   M30xTrimDeck_xOSR_OpenOnCleaning : BOOL; {access Read Only}
   M30xTrimDeckAutoResetOppOpSide : TIMER[5] := ([0].PRE := 500); {access Read Only}
   M30xTrimDeckAutoResetOppOpSideTimeout : TIMER[5] := ([0].PRE := 2000); {access Read Only}
   M30xTrimDeckAutoResetOpSide : TIMER[5] := ([0].PRE := 500); {access Read Only}
   M30xTrimDeckAutoResetOpSideTimeout : TIMER[5] := ([0].PRE := 2000); {access Read Only}
   M30xTrimDeckDriveErrorOppOpSide : TIMER[5] := ([0].PRE := 800); {access Read Only}
   M30xTrimDeckDriveErrorOpSide : TIMER[5] := ([0].PRE := 800); {access Read Only}
   M30xTrimWheel : MAC_TrimmingWheels[5] := ([0].CONF_dTrimWheelCodeOpt := 1, [0].CONF_dPositionWheel_cmm := 687500, [0].CONF_dConveyorLength_cmm := 914500, [0].CONF_dMaxLengthWorkable_cmm := 610000, [0].CONF_dTolerance_cmm[0] := 200, [0].CONF_dTolerance_cmm[1] := 200, [0].CONF_dTrimWheelArmPos_cmm[0] := 687500, [0].CONF_dTrimWheelArmPos_cmm[1] := 687500, [0].CONF_dMaxTimeToReachPosition_ms[0] := 600, [0].CONF_dMaxTimeToReachPosition_ms[1] := 600, [0].CONF_dTrimWheelPresetZero_cmm[0] := 2620, [0].CONF_dTrimWheelPresetZero_cmm[1] := 2560, [0].CONF_dTrimWheelTargetWindow_cmm[0] := 200, [0].CONF_dTrimWheelTargetWindow_cmm[1] := 200, [0].CONF_dTrimWheelMinPos_cmm[0] := 115000, [0].CONF_dTrimWheelMinPos_cmm[1] := 115000, [0].CONF_dTrimWheelMaxPos_cmm[0] := 262000, [0].CONF_dTrimWheelMaxPos_cmm[1] := 256000, [0].CONF_dTrimWheelMinRange_cmm[0] := 115000, [0].CONF_dTrimWheelMinRange_cmm[1] := 115000, [0].CONF_dTrimWheelMaxRange_cmm[0] := 262000, [0].CONF_dTrimWheelMaxRange_cmm[1] := 256000, [0].CONF_dAutoSpeed_mm_min[0] := 1000, [0].CONF_dAutoSpeed_mm_min[1] := 1000, [0].CONF_dManualSpeed_mm_min[0] := 200, [0].CONF_dManualSpeed_mm_min[1] := 200, [0].CONF_rAcceleration_m_s2[0] := 1.0, [0].CONF_rAcceleration_m_s2[1] := 1.0, [0].CONF_rDeceleration_m_s2[0] := 1.0, [0].CONF_rDeceleration_m_s2[1] := 1.0, [0].ST_xInitialConditionOpSideOK := 1, [0].ST_xInitialConditionOppOpSideOK := 1, [0].ST_xCleaningConditionOK := 1, [0].ST_xConditionOKStopCycle := 1, [0].ST_xOutputEnableOpSide := 1, [0].ST_xOutputEnableOppOpSide := 1, [0].ST_xEnableControlError := 1, [0].ST_xInPositionOpSide := 1, [0].ST_xInPositionOppOpSide := 1, [0].INPUT_xProtectionMotor := 3, [0].INPUT_xLocalSafetySwitch := 3, [0].INPUT_xMotorThermalProbe := 3, [0].INPUT_xProtectionBrake := 3, [0].INPUT_xBrakeFeedback := 3, [0].INPUT_xDriveReady := 3, [0].INPUT_xHomePosition := 3, [0].OUTPUT_xDriveEnable := 3, [0].AUX_dReqLengthPlate_cmm[0] := 260000, [0].AUX_dReqLengthPlate_cmm[1] := 260000, [0].AUX_dReqPositionPlate_cmm[0] := 965963, [0].AUX_dReqPositionPlate_cmm[1] := 965963, [0].AUX_dReqTargetPosTranslation_cmm[0] := 190430, [0].AUX_dReqTargetPosTranslation_cmm[1] := 186570, [0].AUX_dHeadPosition_cmm[0] := 965963, [0].AUX_dHeadPosition_cmm[1] := 965963, [0].AUX_dLengthPlate_cmm[0] := 260000, [0].AUX_dLengthPlate_cmm[1] := 260000, [0].AUX_dPositionWheelBrk_cmm[0] := 188408, [0].AUX_dPositionWheelBrk_cmm[1] := 187480, [0].AUX_dActTransPosition_cmm[0] := 188408,
        [0].AUX_dActTransPosition_cmm[1] := 187480, [0].AUX_dOffsetStep[0] := 500, [0].AUX_dOffsetStep[1] := 500, [0].AUX_dFinalTarget_cmm[0] := 188430, [0].AUX_dFinalTarget_cmm[1] := 187570, [0].AUX_dReqSpeed_mm_min[0] := 1000, [0].AUX_dReqSpeed_mm_min[1] := 1000, [0].AUX_dRealSpeed_mm_min[0] := 1000, [0].AUX_dRealSpeed_mm_min[1] := 1000, [0].AUX_dTotalCaps[0] := 1, [0].AUX_dTotalCaps[1] := 1, [0].AUX_rgxActivate[0] := 2, [0].AUX_rgxActivate[1] := 2, [0].AUX_dSearchPlateDataOpSide.dReaction_cmm := 1000, [0].AUX_dSearchPlateDataOpSide.dPositionDecision_cmm := 647500, [0].AUX_dSearchPlateDataOpSide.dPositionStopSearch_cmm := 686500, [0].AUX_dSearchPlateDataOpSide.dPositionStopHooked_cmm := 706500, [0].AUX_dSearchPlateDataOppOpSide.dReaction_cmm := 1000, [0].AUX_dSearchPlateDataOppOpSide.dPositionDecision_cmm := 647500, [0].AUX_dSearchPlateDataOppOpSide.dPositionStopSearch_cmm := 686500, [0].AUX_dSearchPlateDataOppOpSide.dPositionStopHooked_cmm := 706500, [0].AUX_dSearchPlateDataTranslationOpSide.dReaction_cmm := 1000, [0].AUX_dSearchPlateDataTranslationOpSide.dPositionDecision_cmm := 647500, [0].AUX_dSearchPlateDataTranslationOpSide.dPositionStopSearch_cmm := 686500, [0].AUX_dSearchPlateDataTranslationOpSide.dPositionStopHooked_cmm := 706500, [0].AUX_dSearchPlateDataTranslationOppOpSide.dReaction_cmm := 1000, [0].AUX_dSearchPlateDataTranslationOppOpSide.dPositionDecision_cmm := 647500, [0].AUX_dSearchPlateDataTranslationOppOpSide.dPositionStopSearch_cmm := 686500, [0].AUX_dSearchPlateDataTranslationOppOpSide.dPositionStopHooked_cmm := 706500, [0].tmON_TrimWheelTimeOut[0].PRE := 2500, [0].tmON_TrimWheelTimeOut[1].PRE := 2500, [0].tmON_TrimWheelBlow[0].PRE := 880, [0].tmON_TrimWheelBlow[0].ACC := 880, [0].tmON_TrimWheelBlow[1].PRE := 800, [0].tmON_TrimWheelBlow[1].ACC := 800, [0].tmOF_DriveEnable[0].PRE := 30000, [0].tmOF_DriveEnable[0].ACC := 9881, [0].tmOF_DriveEnable[0].TT := 1, [0].tmOF_DriveEnable[0].DN := 1, [0].tmOF_DriveEnable[1].PRE := 30000, [0].tmOF_DriveEnable[1].ACC := 9881, [0].tmOF_DriveEnable[1].TT := 1, [0].tmOF_DriveEnable[1].DN := 1, [0].tmON_FeedbackTimeOut[0].PRE := 3500, [0].tmON_FeedbackTimeOut[1].PRE := 3500, [0].tmON_FeedbackDriveReady[0].PRE := 1000, [0].tmON_FeedbackDriveReady[1].PRE := 1000, [1].CONF_dTrimWheelCodeOpt := 2, [1].CONF_dPositionWheel_cmm := 924500, [1].CONF_dConveyorLength_cmm := 914500, [1].CONF_dMaxLengthWorkable_cmm := 610000, [1].CONF_dTolerance_cmm[0] := 200, [1].CONF_dTolerance_cmm[1] := 200, [1].CONF_dTrimWheelArmPos_cmm[0] := 924500, [1].CONF_dTrimWheelArmPos_cmm[1] := 924500, [1].CONF_dMaxTimeToReachPosition_ms[0] := 600, [1].CONF_dMaxTimeToReachPosition_ms[1] := 600, [1].CONF_dTrimWheelPresetZero_cmm[0] := 260, [1].CONF_dTrimWheelPresetZero_cmm[1] := 260, [1].CONF_dTrimWheelTargetWindow_cmm[0] := 200,
        [1].CONF_dTrimWheelTargetWindow_cmm[1] := 200, [1].CONF_dTrimWheelMinPos_cmm[0] := -15000, [1].CONF_dTrimWheelMinPos_cmm[1] := -15000, [1].CONF_dTrimWheelMaxPos_cmm[0] := 42000, [1].CONF_dTrimWheelMaxPos_cmm[1] := 42000, [1].CONF_dTrimWheelMinRange_cmm[0] := -15000, [1].CONF_dTrimWheelMinRange_cmm[1] := -15000, [1].CONF_dTrimWheelMaxRange_cmm[0] := 42000, [1].CONF_dTrimWheelMaxRange_cmm[1] := 42000, [1].CONF_dAutoSpeed_mm_min[0] := 1000, [1].CONF_dAutoSpeed_mm_min[1] := 1000, [1].CONF_dManualSpeed_mm_min[0] := 200, [1].CONF_dManualSpeed_mm_min[1] := 200, [1].CONF_rAcceleration_m_s2[0] := 1.0, [1].CONF_rAcceleration_m_s2[1] := 1.0, [1].CONF_rDeceleration_m_s2[0] := 1.0, [1].CONF_rDeceleration_m_s2[1] := 1.0, [1].ST_xTailBreakOppOpSide := 1, [1].ST_xInitialConditionOpSideOK := 1, [1].ST_xInitialConditionOppOpSideOK := 1, [1].ST_xCleaningConditionOK := 1, [1].ST_xConditionOKStopCycle := 1, [1].ST_xOutputEnableOpSide := 1, [1].ST_xOutputEnableOppOpSide := 1, [1].ST_xEnableControlError := 1, [1].ST_xInPositionOpSide := 1, [1].ST_xInPositionOppOpSide := 1, [1].ST_xTailBreakOpSide := 1, [1].INPUT_xProtectionMotor := 3, [1].INPUT_xLocalSafetySwitch := 3, [1].INPUT_xMotorThermalProbe := 3, [1].INPUT_xProtectionBrake := 3, [1].INPUT_xBrakeFeedback := 3, [1].INPUT_xDriveReady := 3, [1].INPUT_xHomePosition := 3, [1].OUTPUT_xDriveEnable := 3, [1].AUX_dReqLengthPlate_cmm[0] := 260000, [1].AUX_dReqLengthPlate_cmm[1] := 260000, [1].AUX_dReqPositionPlate_cmm[0] := 1192693, [1].AUX_dReqPositionPlate_cmm[1] := 1192693, [1].AUX_dHeadPosition_cmm[0] := 932693, [1].AUX_dHeadPosition_cmm[1] := 932693, [1].AUX_dPositionWheelBrk_cmm[0] := 13982, [1].AUX_dPositionWheelBrk_cmm[1] := -2494, [1].AUX_dDifferPositionBrkTailMode_cmm[0] := 260000, [1].AUX_dDifferPositionBrkTailMode_cmm[1] := 260000, [1].AUX_dActTransPosition_cmm[0] := 13982, [1].AUX_dActTransPosition_cmm[1] := -2494, [1].AUX_dOffsetStep[0] := 500, [1].AUX_dOffsetStep[1] := 500, [1].AUX_dFinalTarget_cmm[0] := 14000, [1].AUX_dFinalTarget_cmm[1] := -2500, [1].AUX_dReqSpeed_mm_min[0] := 1000, [1].AUX_dReqSpeed_mm_min[1] := 1000, [1].AUX_dRealSpeed_mm_min[0] := 1000, [1].AUX_dRealSpeed_mm_min[1] := 1000, [1].AUX_dTotalCaps[0] := 1, [1].AUX_dTotalCaps[1] := 1, [1].AUX_dSearchPlateDataOpSide.dReaction_cmm := 1000, [1].AUX_dSearchPlateDataOpSide.dPositionDecision_cmm := 914500,
        [1].AUX_dSearchPlateDataOpSide.dPositionStopSearch_cmm := 923500, [1].AUX_dSearchPlateDataOpSide.dPositionStopHooked_cmm := 933500, [1].AUX_dSearchPlateDataOppOpSide.dReaction_cmm := 1000, [1].AUX_dSearchPlateDataOppOpSide.dPositionDecision_cmm := 914500, [1].AUX_dSearchPlateDataOppOpSide.dPositionStopSearch_cmm := 923500, [1].AUX_dSearchPlateDataOppOpSide.dPositionStopHooked_cmm := 933500, [1].AUX_dSearchPlateDataTranslationOpSide.dReaction_cmm := 1000, [1].AUX_dSearchPlateDataTranslationOpSide.dPositionDecision_cmm := 884500, [1].AUX_dSearchPlateDataTranslationOpSide.dPositionStopSearch_cmm := 923500, [1].AUX_dSearchPlateDataTranslationOpSide.dPositionStopHooked_cmm := 943500, [1].AUX_dSearchPlateDataTranslationOppOpSide.dReaction_cmm := 1000, [1].AUX_dSearchPlateDataTranslationOppOpSide.dPositionDecision_cmm := 884500, [1].AUX_dSearchPlateDataTranslationOppOpSide.dPositionStopSearch_cmm := 923500, [1].AUX_dSearchPlateDataTranslationOppOpSide.dPositionStopHooked_cmm := 943500, [1].tmON_TrimWheelTimeOut[0].PRE := 2500, [1].tmON_TrimWheelTimeOut[1].PRE := 2500, [1].tmON_TrimWheelBlow[0].PRE := 500, [1].tmON_TrimWheelBlow[0].ACC := 500, [1].tmON_TrimWheelBlow[1].PRE := 500, [1].tmON_TrimWheelBlow[1].ACC := 500, [1].tmOF_DriveEnable[0].PRE := 30000, [1].tmOF_DriveEnable[0].ACC := 6041, [1].tmOF_DriveEnable[0].TT := 1, [1].tmOF_DriveEnable[0].DN := 1, [1].tmOF_DriveEnable[1].PRE := 30000, [1].tmOF_DriveEnable[1].ACC := 6041, [1].tmOF_DriveEnable[1].TT := 1, [1].tmOF_DriveEnable[1].DN := 1, [1].tmON_FeedbackTimeOut[0].PRE := 3500, [1].tmON_FeedbackTimeOut[1].PRE := 3500, [1].tmON_FeedbackDriveReady[0].PRE := 1000, [1].tmON_FeedbackDriveReady[1].PRE := 1000, [2].CONF_dTrimWheelCodeOpt := 3, [2].CONF_dPositionWheel_cmm := 1432500, [2].CONF_dConveyorLength_cmm := 914500, [2].CONF_dMaxLengthWorkable_cmm := 610000, [2].CONF_dTolerance_cmm[0] := 200, [2].CONF_dTolerance_cmm[1] := 200, [2].CONF_dTrimWheelArmPos_cmm[0] := 1432500, [2].CONF_dTrimWheelArmPos_cmm[1] := 1432500, [2].CONF_dMaxTimeToReachPosition_ms[0] := 600, [2].CONF_dMaxTimeToReachPosition_ms[1] := 600, [2].CONF_dTrimWheelPresetZero_cmm[0] := 260, [2].CONF_dTrimWheelPresetZero_cmm[1] := 260, [2].CONF_dTrimWheelTargetWindow_cmm[0] := 200, [2].CONF_dTrimWheelTargetWindow_cmm[1] := 200, [2].CONF_dTrimWheelMinPos_cmm[0] := -15000, [2].CONF_dTrimWheelMinPos_cmm[1] := -15000, [2].CONF_dTrimWheelMaxPos_cmm[0] := 42000, [2].CONF_dTrimWheelMaxPos_cmm[1] := 42000, [2].CONF_dTrimWheelMinRange_cmm[0] := -15000, [2].CONF_dTrimWheelMinRange_cmm[1] := -15000, [2].CONF_dTrimWheelMaxRange_cmm[0] := 42000, [2].CONF_dTrimWheelMaxRange_cmm[1] := 42000, [2].CONF_dAutoSpeed_mm_min[0] := 1000, [2].CONF_dAutoSpeed_mm_min[1] := 1000, [2].CONF_dManualSpeed_mm_min[0] := 200, [2].CONF_dManualSpeed_mm_min[1] := 200, [2].CONF_rAcceleration_m_s2[0] := 1.0, [2].CONF_rAcceleration_m_s2[1] := 1.0,
        [2].CONF_rDeceleration_m_s2[0] := 1.0, [2].CONF_rDeceleration_m_s2[1] := 1.0, [2].ST_xInitialConditionOpSideOK := 1, [2].ST_xInitialConditionOppOpSideOK := 1, [2].ST_xCleaningConditionOK := 1, [2].ST_xConditionOKStopCycle := 1, [2].ST_xOutputEnableOpSide := 1, [2].ST_xOutputEnableOppOpSide := 1, [2].ST_xEnableControlError := 1, [2].ST_xInPositionOpSide := 1, [2].ST_xInPositionOppOpSide := 1, [2].INPUT_xProtectionMotor := 3, [2].INPUT_xLocalSafetySwitch := 3, [2].INPUT_xMotorThermalProbe := 3, [2].INPUT_xProtectionBrake := 3, [2].INPUT_xBrakeFeedback := 3, [2].INPUT_xDriveReady := 3, [2].INPUT_xHomePosition := 3, [2].OUTPUT_xDriveEnable := 3, [2].AUX_dReqLengthPlate_cmm[0] := 260000, [2].AUX_dReqLengthPlate_cmm[1] := 260000, [2].AUX_dReqPositionPlate_cmm[0] := 1711214, [2].AUX_dReqPositionPlate_cmm[1] := 1711214, [2].AUX_dHeadPosition_cmm[0] := 1711214, [2].AUX_dHeadPosition_cmm[1] := 1711214, [2].AUX_dLengthPlate_cmm[0] := 260000, [2].AUX_dLengthPlate_cmm[1] := 260000, [2].AUX_dPositionWheelBrk_cmm[0] := 484, [2].AUX_dPositionWheelBrk_cmm[1] := -1003, [2].AUX_dActTransPosition_cmm[0] := 484, [2].AUX_dActTransPosition_cmm[1] := -1003, [2].AUX_dOffsetStep[0] := 500, [2].AUX_dOffsetStep[1] := 500, [2].AUX_dFinalTarget_cmm[0] := 500, [2].AUX_dFinalTarget_cmm[1] := -1000, [2].AUX_dReqSpeed_mm_min[0] := 1000, [2].AUX_dReqSpeed_mm_min[1] := 1000, [2].AUX_dRealSpeed_mm_min[0] := 1000, [2].AUX_dRealSpeed_mm_min[1] := 1000, [2].AUX_dTotalCaps[0] := 1, [2].AUX_dTotalCaps[1] := 1, [2].AUX_rgxActivate[0] := 2, [2].AUX_rgxActivate[1] := 2, [2].AUX_dSearchPlateDataOpSide.dReaction_cmm := 1000, [2].AUX_dSearchPlateDataOpSide.dPositionDecision_cmm := 1392500, [2].AUX_dSearchPlateDataOpSide.dPositionStopSearch_cmm := 1431500, [2].AUX_dSearchPlateDataOpSide.dPositionStopHooked_cmm := 1451500, [2].AUX_dSearchPlateDataOppOpSide.dReaction_cmm := 1000, [2].AUX_dSearchPlateDataOppOpSide.dPositionDecision_cmm := 1392500, [2].AUX_dSearchPlateDataOppOpSide.dPositionStopSearch_cmm := 1431500, [2].AUX_dSearchPlateDataOppOpSide.dPositionStopHooked_cmm := 1451500, [2].AUX_dSearchPlateDataTranslationOpSide.dReaction_cmm := 1000, [2].AUX_dSearchPlateDataTranslationOpSide.dPositionDecision_cmm := 1392500, [2].AUX_dSearchPlateDataTranslationOpSide.dPositionStopSearch_cmm := 1431500, [2].AUX_dSearchPlateDataTranslationOpSide.dPositionStopHooked_cmm := 1451500, [2].AUX_dSearchPlateDataTranslationOppOpSide.dReaction_cmm := 1000, [2].AUX_dSearchPlateDataTranslationOppOpSide.dPositionDecision_cmm := 1392500, [2].AUX_dSearchPlateDataTranslationOppOpSide.dPositionStopSearch_cmm := 1431500, [2].AUX_dSearchPlateDataTranslationOppOpSide.dPositionStopHooked_cmm := 1451500, [2].tmON_TrimWheelTimeOut[0].PRE := 2500,
        [2].tmON_TrimWheelTimeOut[1].PRE := 2500, [2].tmON_TrimWheelBlow[0].PRE := 2000, [2].tmON_TrimWheelBlow[0].ACC := 2000, [2].tmON_TrimWheelBlow[1].PRE := 2000, [2].tmON_TrimWheelBlow[1].ACC := 2000, [2].tmOF_DriveEnable[0].PRE := 30000, [2].tmOF_DriveEnable[0].ACC := 12181, [2].tmOF_DriveEnable[0].TT := 1, [2].tmOF_DriveEnable[0].DN := 1, [2].tmOF_DriveEnable[1].PRE := 30000, [2].tmOF_DriveEnable[1].ACC := 12181, [2].tmOF_DriveEnable[1].TT := 1, [2].tmOF_DriveEnable[1].DN := 1, [2].tmON_FeedbackTimeOut[0].PRE := 3500, [2].tmON_FeedbackTimeOut[1].PRE := 3500, [2].tmON_FeedbackDriveReady[0].PRE := 1000, [2].tmON_FeedbackDriveReady[1].PRE := 1000, [3].CONF_dTrimWheelCodeOpt := 4, [3].CONF_dPositionWheel_cmm := 1452500, [3].CONF_dConveyorLength_cmm := 914500, [3].CONF_dMaxLengthWorkable_cmm := 610000, [3].CONF_dTolerance_cmm[0] := 200, [3].CONF_dTolerance_cmm[1] := 200, [3].CONF_dTrimWheelArmPos_cmm[0] := 1452500, [3].CONF_dTrimWheelArmPos_cmm[1] := 1452500, [3].CONF_dMaxTimeToReachPosition_ms[0] := 600, [3].CONF_dMaxTimeToReachPosition_ms[1] := 600, [3].CONF_dTrimWheelPresetZero_cmm[0] := 260, [3].CONF_dTrimWheelPresetZero_cmm[1] := 260, [3].CONF_dTrimWheelTargetWindow_cmm[0] := 200, [3].CONF_dTrimWheelTargetWindow_cmm[1] := 200, [3].CONF_dTrimWheelMinPos_cmm[0] := -15000, [3].CONF_dTrimWheelMinPos_cmm[1] := -15000, [3].CONF_dTrimWheelMaxPos_cmm[0] := 42000, [3].CONF_dTrimWheelMaxPos_cmm[1] := 42000, [3].CONF_dTrimWheelMinRange_cmm[0] := -15000, [3].CONF_dTrimWheelMinRange_cmm[1] := -15000, [3].CONF_dTrimWheelMaxRange_cmm[0] := 42000, [3].CONF_dTrimWheelMaxRange_cmm[1] := 42000, [3].CONF_dAutoSpeed_mm_min[0] := 1000, [3].CONF_dAutoSpeed_mm_min[1] := 1000, [3].CONF_dManualSpeed_mm_min[0] := 200, [3].CONF_dManualSpeed_mm_min[1] := 200, [3].CONF_rAcceleration_m_s2[0] := 1.0, [3].CONF_rAcceleration_m_s2[1] := 1.0, [3].CONF_rDeceleration_m_s2[0] := 1.0, [3].CONF_rDeceleration_m_s2[1] := 1.0, [3].ST_xInitialConditionOpSideOK := 1, [3].ST_xInitialConditionOppOpSideOK := 1, [3].ST_xCleaningConditionOK := 1, [3].ST_xConditionOKStopCycle := 1, [3].ST_xOutputEnableOpSide := 1, [3].ST_xOutputEnableOppOpSide := 1, [3].ST_xEnableControlError := 1, [3].ST_xInPositionOpSide := 1, [3].ST_xInPositionOppOpSide := 1, [3].INPUT_xProtectionMotor := 3, [3].INPUT_xLocalSafetySwitch := 3, [3].INPUT_xMotorThermalProbe := 3, [3].INPUT_xProtectionBrake := 3,
        [3].INPUT_xBrakeFeedback := 3, [3].INPUT_xDriveReady := 3, [3].INPUT_xHomePosition := 3, [3].OUTPUT_xDriveEnable := 3, [3].AUX_dReqLengthPlate_cmm[0] := 260000, [3].AUX_dReqLengthPlate_cmm[1] := 260000, [3].AUX_dReqPositionPlate_cmm[0] := 1730648, [3].AUX_dReqPositionPlate_cmm[1] := 1730648, [3].AUX_dHeadPosition_cmm[0] := 1730648, [3].AUX_dHeadPosition_cmm[1] := 1730648, [3].AUX_dPositionWheelBrk_cmm[0] := -503, [3].AUX_dPositionWheelBrk_cmm[1] := 3, [3].AUX_dActTransPosition_cmm[0] := -503, [3].AUX_dActTransPosition_cmm[1] := 3, [3].AUX_dOffsetStep[0] := 500, [3].AUX_dOffsetStep[1] := 500, [3].AUX_dFinalTarget_cmm[0] := -500, [3].AUX_dReqSpeed_mm_min[0] := 1000, [3].AUX_dReqSpeed_mm_min[1] := 1000, [3].AUX_dRealSpeed_mm_min[0] := 1000, [3].AUX_dRealSpeed_mm_min[1] := 1000, [3].AUX_dTotalCaps[0] := 1, [3].AUX_dTotalCaps[1] := 1, [3].AUX_rgxActivate[0] := 2, [3].AUX_rgxActivate[1] := 2, [3].AUX_dSearchPlateDataOpSide.dReaction_cmm := 1000, [3].AUX_dSearchPlateDataOpSide.dPositionDecision_cmm := 1412500, [3].AUX_dSearchPlateDataOpSide.dPositionStopSearch_cmm := 1451500, [3].AUX_dSearchPlateDataOpSide.dPositionStopHooked_cmm := 1471500, [3].AUX_dSearchPlateDataOppOpSide.dReaction_cmm := 1000, [3].AUX_dSearchPlateDataOppOpSide.dPositionDecision_cmm := 1412500, [3].AUX_dSearchPlateDataOppOpSide.dPositionStopSearch_cmm := 1451500, [3].AUX_dSearchPlateDataOppOpSide.dPositionStopHooked_cmm := 1471500, [3].AUX_dSearchPlateDataTranslationOpSide.dReaction_cmm := 1000, [3].AUX_dSearchPlateDataTranslationOpSide.dPositionDecision_cmm := 1412500, [3].AUX_dSearchPlateDataTranslationOpSide.dPositionStopSearch_cmm := 1451500, [3].AUX_dSearchPlateDataTranslationOpSide.dPositionStopHooked_cmm := 1471500, [3].AUX_dSearchPlateDataTranslationOppOpSide.dReaction_cmm := 1000, [3].AUX_dSearchPlateDataTranslationOppOpSide.dPositionDecision_cmm := 1412500, [3].AUX_dSearchPlateDataTranslationOppOpSide.dPositionStopSearch_cmm := 1451500, [3].AUX_dSearchPlateDataTranslationOppOpSide.dPositionStopHooked_cmm := 1471500, [3].tmON_TrimWheelTimeOut[0].PRE := 2500, [3].tmON_TrimWheelTimeOut[1].PRE := 2500, [3].tmON_TrimWheelBlow[0].PRE := 500, [3].tmON_TrimWheelBlow[0].ACC := 501, [3].tmON_TrimWheelBlow[1].PRE := 500, [3].tmON_TrimWheelBlow[1].ACC := 501, [3].tmOF_DriveEnable[0].PRE := 30000, [3].tmOF_DriveEnable[0].ACC := 11901, [3].tmOF_DriveEnable[0].TT := 1, [3].tmOF_DriveEnable[0].DN := 1, [3].tmOF_DriveEnable[1].PRE := 30000, [3].tmOF_DriveEnable[1].ACC := 11901, [3].tmOF_DriveEnable[1].TT := 1, [3].tmOF_DriveEnable[1].DN := 1, [3].tmON_FeedbackTimeOut[0].PRE := 3500, [3].tmON_FeedbackTimeOut[1].PRE := 3500, [3].tmON_FeedbackDriveReady[0].PRE := 1000, [3].tmON_FeedbackDriveReady[1].PRE := 1000); {access None}
        [2]   // M303C1
        [3]   // M303C2
        [0]   // M303A
        [1]   // M303B
   M30xTrimWheel_ALM : MAC_TrimmingWheels_ALM[5]; {access Read Only}
        [0].rgxStoppingFault[0].x11   // M302.Trimming wheel drive error opposite operator side
        [0].rgxStoppingFault[0].x12   // M302.Trimming wheel drive feedback error opposite operator side
        [0].rgxStoppingFault[0].x14   // M302.Trimming wheel feedback brake opposite operator side
        [1].rgxStoppingFault[0].x14   // M303.Trimming wheel feedback brake opposite operator side
        [0].rgxStoppingFault[0].x2   // M302.Trimming wheel drive feedback error operator side
        [0].rgxStoppingFault[0].x10   // M302.Trimming wheel protection motor opposite operator side
        [0].rgxStoppingFault[0].x13   // M302.Trimming wheel protection brake opposite operator side
        [1].rgxStoppingFault[0].x11   // M303.Trimming wheel drive error opposite operator side
        [1].rgxStoppingFault[0].x12   // M303.Trimming wheel drive feedback error opposite operator side
        [2]   // M304
        [0]   // M302
        [3]   // M305
        [1]   // M303
        [0].rgxStoppingFault[0].x6   // M302.Drive not enabled operator side
        [0].rgxStoppingFault[0].x1   // M302.Trimming wheel drive error operator side
        [0].rgxStoppingFault[0].x15   // M302.Motor thermal probe opposite operator side
        [0].rgxStoppingFault[0].x4   // M302.Trimming wheel feedback brake operator side
        [0].rgxStoppingFault[0].x16   // M302.Drive not enabled opposite operator side
        [0].rgxStoppingFault[0].x3   // M302.Trimming wheel protection brake operator side
        [0].rgxStoppingFault[0].x0   // M302.Trimming wheel protection motor operator side
        [0].rgxStoppingFault[0].x5   // M302.Motor thermal probe operator side
        [0].rgxFault[0].x10   // M302.Trimming wheel position error opposite operator side
        [0].rgxFault[0].x0   // M302.Trimming wheel position error operator side
        [1].rgxStoppingFault[0].x6   // M303.Drive not enabled operator side
        [1].rgxStoppingFault[0].x2   // M303.Trimming wheel drive feedback error operator side
        [1].rgxStoppingFault[0].x10   // M303.Trimming wheel protection motor opposite operator side
        [1].rgxStoppingFault[0].x1   // M303.Trimming wheel drive error operator side
        [1].rgxStoppingFault[0].x15   // M303.Motor thermal probe opposite operator side
        [1].rgxStoppingFault[0].x13   // M303.Trimming wheel protection brake opposite operator side
        [1].rgxStoppingFault[0].x4   // M303.Trimming wheel feedback brake operator side
        [1].rgxStoppingFault[0].x16   // M303.Drive not enabled opposite operator side
        [1].rgxStoppingFault[0].x3   // M303.Trimming wheel protection brake operator side
        [1].rgxStoppingFault[0].x0   // M303.Trimming wheel protection motor operator side
        [1].rgxStoppingFault[0].x5   // M303.Motor thermal probe operator side
        [1].rgxFault[0].x10   // M303.Trimming wheel position error opposite operator side
        [1].rgxFault[0].x0   // M303.Trimming wheel position error operator side
        [2].rgxStoppingFault[0].x11   // M304.Trimming wheel drive error opposite operator side
        [2].rgxStoppingFault[0].x6   // M304.Drive not enabled operator side
        [2].rgxStoppingFault[0].x12   // M304.Trimming wheel drive feedback error opposite operator side
        [2].rgxStoppingFault[0].x14   // M304.Trimming wheel feedback brake opposite operator side
        [2].rgxStoppingFault[0].x2   // M304.Trimming wheel drive feedback error operator side
        [2].rgxStoppingFault[0].x10   // M304.Trimming wheel protection motor opposite operator side
        [2].rgxStoppingFault[0].x1   // M304.Trimming wheel drive error operator side
        [2].rgxStoppingFault[0].x15   // M304.Motor thermal probe opposite operator side
        [2].rgxStoppingFault[0].x13   // M304.Trimming wheel protection brake opposite operator side
        [2].rgxStoppingFault[0].x4   // M304.Trimming wheel feedback brake operator side
        [2].rgxStoppingFault[0].x16   // M304.Drive not enabled opposite operator side
        [2].rgxStoppingFault[0].x3   // M304.Trimming wheel protection brake operator side
        [2].rgxStoppingFault[0].x0   // M304.Trimming wheel protection motor operator side
        [2].rgxStoppingFault[0].x5   // M304.Motor thermal probe operator side
        [2].rgxFault[0].x10   // M304.Trimming wheel position error opposite operator side
        [2].rgxFault[0].x0   // M304.Trimming wheel position error operator side
        [3].rgxStoppingFault[0].x11   // M305.Trimming wheel drive error opposite operator side
        [3].rgxStoppingFault[0].x6   // M305.Drive not enabled operator side
        [3].rgxStoppingFault[0].x12   // M305.Trimming wheel drive feedback error opposite operator side
        [3].rgxStoppingFault[0].x14   // M305.Trimming wheel feedback brake opposite operator side
        [3].rgxStoppingFault[0].x2   // M305.Trimming wheel drive feedback error operator side
        [3].rgxStoppingFault[0].x10   // M305.Trimming wheel protection motor opposite operator side
        [3].rgxStoppingFault[0].x1   // M305.Trimming wheel drive error operator side
        [3].rgxStoppingFault[0].x15   // M305.Motor thermal probe opposite operator side
        [3].rgxStoppingFault[0].x13   // M305.Trimming wheel protection brake opposite operator side
        [3].rgxStoppingFault[0].x4   // M305.Trimming wheel feedback brake operator side
        [3].rgxStoppingFault[0].x16   // M305.Drive not enabled opposite operator side
        [3].rgxStoppingFault[0].x3   // M305.Trimming wheel protection brake operator side
        [3].rgxStoppingFault[0].x0   // M305.Trimming wheel protection motor operator side
        [3].rgxStoppingFault[0].x5   // M305.Motor thermal probe operator side
        [3].rgxFault[0].x10   // M305.Trimming wheel position error opposite operator side
        [3].rgxFault[0].x0   // M305.Trimming wheel position error operator side
        [4]   // M306
        [4].rgxStoppingFault[0].x0   // M306.Trimming wheel protection motor operator side
        [4].rgxStoppingFault[0].x1   // M306.Trimming wheel drive error operator side
        [4].rgxStoppingFault[0].x2   // M306.Trimming wheel drive feedback error operator side
        [4].rgxStoppingFault[0].x3   // M306.Trimming wheel protection brake operator side
        [4].rgxStoppingFault[0].x4   // M306.Trimming wheel feedback brake operator side
        [4].rgxStoppingFault[0].x5   // M306.Motor thermal probe operator side
        [4].rgxStoppingFault[0].x6   // M306.Drive not enabled operator side
        [4].rgxStoppingFault[0].x10   // M306.Trimming wheel protection motor opposite operator side
        [4].rgxStoppingFault[0].x16   // M306.Drive not enabled opposite operator side
        [4].rgxStoppingFault[0].x15   // M306.Motor thermal probe opposite operator side
        [4].rgxStoppingFault[0].x11   // M306.Trimming wheel drive error opposite operator side
        [4].rgxStoppingFault[0].x12   // M306.Trimming wheel drive feedback error opposite operator side
        [4].rgxStoppingFault[0].x13   // M306.Trimming wheel protection brake opposite operator side
        [4].rgxStoppingFault[0].x14   // M306.Trimming wheel feedback brake opposite operator side
        [4].rgxFault[0].x0   // M306.Trimming wheel position error operator side
        [4].rgxFault[0].x10   // M306.Trimming wheel position error opposite operator side
   M30xTrimWheel_DATA : UDT_ConvoyCap_ZC[5];
        [1]   // Cap data M303
        [3]   // Cap data M305
        [0]   // Cap data M302
        [2]   // Cap data M304
        [4]   // Cap data M306
   M30xTrimWheel_HMR : MAC_TrimmingWheels_HMR[5] := ([0].xAutoTrim := 1, [0].xDynamicTrim := 1, [0].xBlowChipsEnabled := 1, [0].xEnabledOpSide := 1, [0].xEnabledOppOpSide := 1, [0].rgdTarget_cmm[0] := 188430, [0].rgdTarget_cmm[1] := 187570, [0].rgdPosition_cmm[0] := 188408, [0].rgdPosition_cmm[1] := 187480, [0].rgdState[0] := 1, [0].rgdState[1] := 1, [1].xAutoTrim := 1, [1].xDynamicTrim := 1, [1].xBlowChipsEnabled := 1, [1].xEnabledOpSide := 1, [1].xEnabledOppOpSide := 1, [1].rgdTarget_cmm[0] := 14000, [1].rgdTarget_cmm[1] := -2500, [1].rgdPosition_cmm[0] := 13982, [1].rgdPosition_cmm[1] := -2494, [1].rgdState[0] := 1, [1].rgdState[1] := 1, [2].xAutoTrim := 1, [2].xDynamicTrim := 1, [2].xBlowChipsEnabled := 1, [2].xEnabledOpSide := 1, [2].xEnabledOppOpSide := 1, [2].xWheelDownOpSide := 1, [2].xWheelDownOppOpSide := 1, [2].rgdTarget_cmm[0] := 500, [2].rgdTarget_cmm[1] := -1000, [2].rgdPosition_cmm[0] := 484, [2].rgdPosition_cmm[1] := -1003, [2].rgdState[0] := 1, [2].rgdState[1] := 1, [3].xAutoTrim := 1, [3].xDynamicTrim := 1, [3].xBlowChipsEnabled := 1, [3].xEnabledOpSide := 1, [3].xEnabledOppOpSide := 1, [3].rgdTarget_cmm[0] := -500, [3].rgdPosition_cmm[0] := -503, [3].rgdPosition_cmm[1] := 3, [3].rgdState[0] := 1, [3].rgdState[1] := 1); {access Read Only}
        [2]   // M304
        [3]   // M305
        [1]   // M303
        [0]   // M302
        [4]   // M306
   M30xTrimWheel_HMW : MAC_TrimmingWheels_HMW[5] := ([0].xEnableDisableBlowChips := 1, [0].rgdBlowTime_ms[0] := 880, [0].rgdBlowTime_ms[1] := 800, [0].rgdOffsetStartTrim_cmm[0] := 30000, [0].rgdOffsetStartTrim_cmm[1] := 30000, [0].rgdReactionTime_ms[0] := 800, [0].rgdReactionTime_ms[1] := 800, [0].rgdOffsetPosition_cmm[0] := -2000, [0].rgdOffsetPosition_cmm[1] := 1000, [0].rgdPlateLengthRise_perc[0] := 100, [0].rgdPlateLengthRise_perc[1] := 100, [1].xEnableDisableBlowChips := 1, [1].rgdBlowTime_ms[0] := 500, [1].rgdBlowTime_ms[1] := 500, [1].rgdOffsetStartTrim_cmm[0] := 25000, [1].rgdOffsetStartTrim_cmm[1] := 40000, [1].rgdOffsetPosition_cmm[0] := 14000, [1].rgdOffsetPosition_cmm[1] := -2500, [1].rgdPlateLengthRise_perc[0] := 100, [1].rgdPlateLengthRise_perc[1] := 100, [2].xEnableDisableBlowChips := 1, [2].rgdBlowTime_ms[0] := 2000, [2].rgdBlowTime_ms[1] := 2000, [2].rgdOffsetStartTrim_cmm[0] := 20000, [2].rgdOffsetStartTrim_cmm[1] := 24000, [2].rgdReactionTime_ms[0] := 800, [2].rgdReactionTime_ms[1] := 800, [2].rgdOffsetPosition_cmm[0] := 500, [2].rgdOffsetPosition_cmm[1] := -1000, [2].rgdPlateLengthRise_perc[0] := 100, [2].rgdPlateLengthRise_perc[1] := 100, [3].xEnableDisableBlowChips := 1, [3].rgdBlowTime_ms[0] := 500, [3].rgdBlowTime_ms[1] := 500, [3].rgdOffsetStartTrim_cmm[0] := 15000, [3].rgdOffsetStartTrim_cmm[1] := 20000, [3].rgdOffsetStopTrim_cmm[0] := -20000, [3].rgdReactionTime_ms[0] := 800, [3].rgdReactionTime_ms[1] := 800, [3].rgdOffsetPosition_cmm[0] := -500, [3].rgdOffsetPosition_cmm[1] := -8500, [3].rgdPlateLengthRise_perc[0] := 100, [3].rgdPlateLengthRise_perc[1] := 100);
        [1]   // M303
        [0]   // M302
        [2]   // M304
        [3]   // M305
        [4]   // M306
   M310_M1_DR_R1 : AXIS_CIP_DRIVE; {access Read Only}
   M310_M2_DR_R2 : AXIS_CIP_DRIVE; {access Read Only}
   M310_M3_DR_R3 : AXIS_CIP_DRIVE; {access Read Only}
   M310_M4_DR_B1 : AXIS_CIP_DRIVE; {access Read Only}
   M310_M5_DR_B2 : AXIS_CIP_DRIVE; {access Read Only}
   M310_M6_DR_L1 : AXIS_CIP_DRIVE; {access Read Only}
   M310_M7_DR_L2 : AXIS_CIP_DRIVE; {access Read Only}
   M310_xReqStopPrevConvForPos : BOOL; {access Read Only}
   M310B : MAC_Conveyor := (ST_xCleaningConditionOK := 1, ST_xConditionOKStopCycle := 1, ST_xEnableControlError := 1, ST_xSafetyMovement := 1, ST_xAux4 := 1, OSR_xSynchroPhotocellTail := 1, INPUT_xLowPositionPopup_1 := 1, INPUT_xLowPositionPopup_2 := 1, INPUT_xDriveReady_M2 := 1, INPUT_xDriveReady_M3 := 1, INPUT_xLocalSafetySwitch_M3 := 1, INPUT_xProtectionMotor_M3 := 1, INPUT_xDriveReady_M4 := 1, INPUT_xLocalSafetySwitch_M4 := 1, INPUT_xProtectionMotor_M4 := 1, OUTPUT_xDriveEnable_M3 := 1, OUTPUT_xDriveEnable_M4 := 1, AUX_dPresetStopLoad_cmm := 455000, AUX_dPresetStopUnload_cmm := 575000, AUX_dAccSpace_cmm := 41667, AUX_dDecSpace_cmm := 41667, AUX_dReqSpeed_mm_min := 60000, AUX_dPhPosTarget_cmm := 180000, TmON_AxleReadyToMoveDelayed.PRE := 500, tmON_FeedbackTimeOut_M1.PRE := 1500, tmOF_DriveEnable_M1.PRE := 20000, tmOF_DriveEnable_M1.ACC := 6500, tmOF_DriveEnable_M1.TT := 1, tmOF_DriveEnable_M1.DN := 1, tmOF_PowerSaving_M1.PRE := 20000, tmOF_PowerSaving_M1.ACC := 20000, tmOF_PowerSaving_M1.EN := 1, tmOF_PowerSaving_M1.DN := 1, tmON_FeedbackTimeOut_M2.PRE := 1500, tmOF_DriveEnable_M2.PRE := 20000, tmOF_DriveEnable_M2.ACC := 3500, tmOF_PowerSaving_M2.PRE := 20000, tmON_FeedbackTimeOut_M3.PRE := 1500, tmOF_DriveEnable_M3.PRE := 20000, tmOF_DriveEnable_M3.ACC := 6500, tmOF_DriveEnable_M3.TT := 1, tmOF_DriveEnable_M3.DN := 1, tmOF_PowerSaving_M3.PRE := 20000, tmOF_PowerSaving_M3.ACC := 20000, tmON_FeedbackTimeOut_M4.PRE := 1500, tmOF_DriveEnable_M4.PRE := 20000, tmOF_DriveEnable_M4.ACC := 3500, tmOF_DriveEnable_M4.TT := 1, tmOF_DriveEnable_M4.DN := 1, tmOF_MCD_M1.PRE := 200, tmOF_MCD_M1.ACC := 200, tmOF_MCD_M2.PRE := 200, tmOF_MCD_M2.ACC := 200, tmOF_MCD_M3.PRE := 200, tmOF_MCD_M3.ACC := 200, tmOF_MCD_M4.PRE := 200, tmOF_MCD_M4.ACC := 200); {access None}
        .INPUT_xMotorThermalProbe_M1   // M310B.M1.P403BT1.Motor thermal probe
        .PH_x.0   // Load
        .PH_x.1   // Load Upstream
        .PH_x.10   // Unload Downstream
        .PH_x.13   // End unload Upstream
        .PH_x.14   // End unload Downstream
        .PH_x.15   // End unload
        .PH_x.16   // Unpack convoy
        .PH_x.17   // End unpack convoy
        .PH_x.18   // Unpack convoy Upstream
        .PH_x.19   // End unpack convoy Upstream
        .PH_x.2   // Load Downstream
        .PH_x.20   // Unpack convoy Downstream
        .PH_x.21   // End unpack convoy Downstream
        .PH_x.22   // Stop for unload on main line
        .PH_x.23   // End stop for unload on main line
        .PH_x.24   // Stop for unload on main line Upstream
        .PH_x.25   // End stop for unload on main line Upstream
        .PH_x.26   // Stop for unload on main line Downstream
        .PH_x.27   // End stop for unload on main line Downstream
        .PH_x.28   // Load reentry
        .PH_x.29   // End load reentry
        .PH_x.5   // End load Upstream
        .PH_x.6   // End load Downstream
        .PH_x.7   // End load
        .PH_x.8   // Unload
        .PH_x.9   // Unload Upstream
        .INPUT_xMotorThermalProbe_M2   // M310B.M2.P403BT2.Motor thermal probe
   M310B_ALM : MAC_Conveyor_ALM;
        .rgxStoppingFault_M[0].13   // Z401.M310B-M2.P51AZ1.Local safety switch
        .rgxStoppingFault_M[0].2   // Z401.M310B-M1.P51AZ1.Drive feedback error
        .rgxStoppingFault_M[0].0   // Z401.M310B-M1.P51AZ1.Protection motor rotation
        .rgxStoppingFault_M[0].4   // Z401.M310B-M1.P403BT1.Motor thermal probe
        .rgxStoppingFault_M[0].12   // Z401.M310B-M2.P51AZ1.Drive feedback error
        .rgxStoppingFault[0].0   // Z401.M310B.Positioning error
        .rgxStoppingFault_M[0].1   // Z401.M310B-M1.P51AZ1.Drive error
        .rgxStoppingFault_M[0].11   // Z401.M310B-M2.P51AZ1.Drive error
        .rgxStoppingFault_M[0].15   // Z401.M310B-M2.P51AZ1.Braking resistor anomaly
        .rgxStoppingFault_M[0].6   // Z401.M310B-M1.Drive not ready
        .rgdFaultCode_M[0]   // Drive fault code M1
        .rgdFaultCode_M[1]   // Drive fault code M2
        .rgxStoppingFault_M[0].5   // Z401.M310B-M1.P51AZ1.Braking resistor anomaly
        .rgxStoppingFault_M[0].16   // Z401.M310B-M2.Drive not ready
        .rgxWarning[0].0   // Z401.M310B.Plate not synchronized
        .rgxStoppingFault_M[0].3   // Z401.M310B-M1.P51AZ1.Local safety switch
        .rgxStoppingFault_M[0].14   // Z401.M310B-M2.P403BT2.Motor thermal probe
        .rgxStoppingFault_M[0].10   // Z401.M310B-M2.P51AZ1.Protection motor rotation
   M310B_Data : UDT_Convoy_SL; {access Read Only}
   M310B_HMR : MAC_Conveyor_HMR := (dState1 := 1, dState3 := 1, dState4 := 1, dStateSensor1 := 1, dStateSensor2 := 1);
        .rgxMan.6   // Run M4 (NU)
        .rgxMan.7   // Reverse M4 (NU)
        .dErrorCode1   // Error code M1
        .rgxMan.0   // Run M1
        .rgxMan.1   // Reverse M1
        .rgxMan.2   // Run M2
        .rgxMan.3   // Reverse M2
        .rgxMan.8   // Run both
        .rgxMan.9   // Reverse both
        .dErrorCode2   // Error code M2
        .dErrorCode4   // Error code M4 (NU)
        .dErrorCode3   // Error code M3 (NU)
        .rgxMan.5   // Reverse M3 (NU)
        .rgxMan.4   // Run M3 (NU)
   M310B_HMW : MAC_Conveyor_HMW;
        .rgxMan.7   // Reverse M4 (NU)
        .rgxMan.5   // Reverse M3 (NU)
        .rgxMan.0   // Run M1
        .rgxMan.1   // Reverse M1
        .rgxMan.2   // Run M2
        .rgxMan.3   // Reverse M2
        .rgxMan.4   // Run M3 (NU)
        .rgxMan.6   // Run M4 (NU)
        .rgxMan.8   // Run both
        .rgxMan.9   // Reverse both
   M310B_M1_DR_IN_MAJ : MOTION_INSTRUCTION := (FLAGS := 570425344, DN := 1); {access None}
   M310B_M1_DR_IN_MAM : MOTION_INSTRUCTION := (FLAGS := 33554432); {access None}
   M310B_M1_DR_IN_MAR : MOTION_INSTRUCTION := (FLAGS := 33554432); {access None}
   M310B_M1_DR_IN_MAS : MOTION_INSTRUCTION := (FLAGS := -1442840576, EN := 1, DN := 1, PC := 1); {access None}
   M310B_M1_DR_IN_MCD : MOTION_INSTRUCTION := (FLAGS := 570425344, DN := 1); {access None}
   M310B_M1_DR_IN_MRP : MOTION_INSTRUCTION := (FLAGS := 33554432); {access None}
   M310B_M1_DR_MAFR : MOTION_INSTRUCTION := (FLAGS := 301989888, ER := 1, ERR := 11); {access None}
   M310B_M1_DR_MDR : MOTION_INSTRUCTION := (FLAGS := -1845493760, EN := 1, ER := 1, ERR := 11); {access None}
   M310B_M1_DR_MSF : MOTION_INSTRUCTION := (FLAGS := 570425344, DN := 1, STATUS := 2, STATE := 1); {access None}
   M310B_M1_DR_MSO : MOTION_INSTRUCTION := (FLAGS := -1610612736, EN := 1, DN := 1, STATE := 1); {access None}
   M310B_M1_DR_OUT_MAJ : MOTION_INSTRUCTION := (FLAGS := 570425344, DN := 1); {access None}
   M310B_M1_DR_OUT_MAM : MOTION_INSTRUCTION := (FLAGS := 33554432); {access None}
   M310B_M1_DR_OUT_MAR : MOTION_INSTRUCTION := (FLAGS := 33554432); {access None}
   M310B_M1_DR_OUT_MAS : MOTION_INSTRUCTION := (FLAGS := -1442840576, EN := 1, DN := 1, PC := 1); {access None}
   M310B_M1_DR_OUT_MCD : MOTION_INSTRUCTION := (FLAGS := 570425344, DN := 1); {access None}
   M310B_M1_DR_OUT_MRP : MOTION_INSTRUCTION := (FLAGS := 33554432); {access None}
   M310B_M2_DR_IN_MAJ : MOTION_INSTRUCTION := (FLAGS := 570425344, DN := 1); {access None}
   M310B_M2_DR_IN_MAM : MOTION_INSTRUCTION := (FLAGS := 33554432); {access None}
   M310B_M2_DR_IN_MAR : MOTION_INSTRUCTION := (FLAGS := 33554432); {access None}
   M310B_M2_DR_IN_MAS : MOTION_INSTRUCTION := (FLAGS := -1442840576, EN := 1, DN := 1, PC := 1); {access None}
   M310B_M2_DR_IN_MCD : MOTION_INSTRUCTION := (FLAGS := 570425344, DN := 1); {access None}
   M310B_M2_DR_IN_MRP : MOTION_INSTRUCTION := (FLAGS := 33554432); {access None}
   M310B_M2_DR_MAFR : MOTION_INSTRUCTION := (FLAGS := 301989888, ER := 1, ERR := 11); {access None}
   M310B_M2_DR_MDR : MOTION_INSTRUCTION := (FLAGS := -1845493760, EN := 1, ER := 1, ERR := 11); {access None}
   M310B_M2_DR_MSF : MOTION_INSTRUCTION := (FLAGS := 570425344, DN := 1, STATUS := 2, STATE := 1); {access None}
   M310B_M2_DR_MSO : MOTION_INSTRUCTION := (FLAGS := -1610612736, EN := 1, DN := 1, STATE := 1); {access None}
   M310B_M2_DR_OUT_MAJ : MOTION_INSTRUCTION := (FLAGS := 570425344, DN := 1); {access None}
   M310B_M2_DR_OUT_MAM : MOTION_INSTRUCTION := (FLAGS := 33554432); {access None}
   M310B_M2_DR_OUT_MAR : MOTION_INSTRUCTION := (FLAGS := 33554432); {access None}
   M310B_M2_DR_OUT_MAS : MOTION_INSTRUCTION := (FLAGS := -1442840576, EN := 1, DN := 1, PC := 1); {access None}
   M310B_M2_DR_OUT_MCD : MOTION_INSTRUCTION := (FLAGS := 570425344, DN := 1); {access None}
   M310B_M2_DR_OUT_MRP : MOTION_INSTRUCTION := (FLAGS := 33554432); {access None}
   M310B_SpaceConv_Utilities : SpaceConv_Utilities := (CONST_dSyncMode := 1, CONST_dSyncroPhWindow_cmm := 450000, CONST_dConveyorLength_cmm := 800000, CONST_dConveyorWidth_cmm := 400000, CONST_dPresetFeedbackTime_ms := 500, CONST_rAcceleration_ms2 := 1.2, CONST_rDeceleration_ms2 := 1.2, CONF_MD1_dScan_ms := 20, CONF_MD2_MD3_dPrstPos_cmm := -390000, CONF_MD4_MD6_dLength_cmm := 365800, CONF_MD7_dOffset_cmm := 50000, ST_dStopLoadForseen_cmm := 620000, ST_dRealSpeed_mm_min := 90000, ST_rStepAdvancementH := 3000.0, ST_rStepAdvancementT := 3000.0, O_xPlateSynchronized := 1, O_dCountFeedbackTime_ms := 500, O_dPresetLoadUnload_cmm := -126300);
   M310B_xOS_PosReq : BOOL;
   M310B_xPlateCullet : BOOL; {access Read Only}
   M310Popup : MAC_Popup_ZC[2] := ([0].ST_xTunnelType := 1, [0].ST_xCleaningConditionOK := 1, [0].ST_xConditionOKForStopCycle := 1, [0].ST_xOutputEnable := 1, [0].ST_xInitialConditionForRise := 1, [0].ST_xExternalConditionToRise := 1, [0].ST_xExternalConditionToDescend := 1, [0].ST_xOutOfEncumbrance := 1, [0].ST_xConditionToReceiveGlass := 1, [0].ST_xEnableControlError := 1, [0].ST_xPlateUnderPopup := 1, [0].ST_xIndexConsPositioning := 1, [0].ST_xPlateComingToPopup := 1, [0].ST_xPlateToBothComing := 1, [0].ST_xPlateToBothPositioning := 1, [0].INPUT_xLiftingProtectionMotor := 1, [0].INPUT_xProtectionCoolingFan := 1, [0].INPUT_xFeedbackCoolingFan := 1, [0].INPUT_xPopupLow := 1, [0].OUTPUT_xPopupVentilation := 1, [0].AUX_dStartPosition_cmm := 4627000, [0].AUX_dEndPosition_cmm := 4827000, [0].AUX_dSpeedConveyor_mm_min := 90000, [0].AUX_dReactionTime_ms := 1500, [0].AUX_dWindowSearch_cmm := 200000, [0].AUX_dDestMaskOpSide := 16#0000_0001, [0].AUX_dReqTarget_cmm := 270000, [0].AUX_dPosPhotocell_cmm := 4627000, [0].AUX_dIndexHead := 3, [0].AUX_dPosTimeout := 5427000, [0].AUX_dIndexPositioning := 3, [0].AUX_dIndexPlateToChangeDestAfterPopup := 1, [0].AUX_tSearchPlateData.dReaction_cmm := 225000, [0].AUX_tSearchPlateData.dPositionDecision_cmm := 4327000, [0].AUX_tSearchPlateData.dPositionStopSearch_cmm := 4627000, [0].AUX_tSearchPlateData.dPositionStopHooked_cmm := 5247000, [0].AUX_tSearchPlateData.dIndex := 3, [0].AUX_tSearchPlateData.xIndexCons := 1, [0].AUX_tSearchPlateData.xPlateHooked := 1, [0].AUX_tSearchPlateData.tResult.rgdHeadPointer[0] := 3, [0].AUX_tSearchPlateData.tResult.rgdHead_cmm[0] := 4328205, [0].AUX_tSearchPlateData.tResult.rgxHead := 1, [0].AUX_tSearchPlateData.tResult.xHeadPresence := 1, [0].tmON_LiftingTimeOut.PRE := 2000, [0].tmON_LiftingFeedbackTimeOut.PRE := 1000, [0].tmOF_WaitBothEndLift.PRE := 1500, [0].tmOF_WaitBothEndLift.ACC := 1500, [0].tmOF_Wait.PRE := 50, [0].tmOF_Wait.ACC := 60, [0].tmON_Saturation.PRE := 1200, [0].tmON_ReentryPlate.PRE := 200, [0].tmON_Positioning.PRE := 40, [1].ST_xTunnelType := 1, [1].ST_xCleaningConditionOK := 1, [1].ST_xConditionOKForStopCycle := 1, [1].ST_xOutputEnable := 1, [1].ST_xInitialConditionForRise := 1, [1].ST_xExternalConditionToRise := 1, [1].ST_xExternalConditionToDescend := 1, [1].ST_xOutOfEncumbrance := 1,
        [1].ST_xConditionToReceiveGlass := 1, [1].ST_xEnableControlError := 1, [1].INPUT_xLiftingProtectionMotor := 1, [1].INPUT_xProtectionCoolingFan := 1, [1].INPUT_xFeedbackCoolingFan := 1, [1].INPUT_xPopupLow := 1, [1].OUTPUT_xPopupVentilation := 1, [1].AUX_dStartPosition_cmm := 4827000, [1].AUX_dEndPosition_cmm := 5027000, [1].AUX_dSpeedConveyor_mm_min := 90000, [1].AUX_dReactionTime_ms := 1500, [1].AUX_dWindowSearch_cmm := 200000, [1].AUX_dDestMaskOpSide := 16#0000_0001, [1].AUX_dPosPhotocell_cmm := 4577000, [1].AUX_dPosTimeout := 5427000, [1].tmON_LiftingTimeOut.PRE := 2000, [1].tmON_LiftingFeedbackTimeOut.PRE := 1000, [1].tmOF_WaitBothEndLift.PRE := 1500, [1].tmOF_WaitBothEndLift.ACC := 1500, [1].tmON_ReentryPlate.PRE := 200, [1].tmON_Positioning.PRE := 40); {access None}
   M310Popup_ALM : MAC_Popup_ZC_ALM[2]; {access Read Only}
        [0].rgxFault[0].0   // M310PopupUP.Lifting protection motor
        [0].rgxFault[0].1   // M310PopupUP.Lifting feedback motor
        [0].rgxFault[0].3   // M310PopupUP.Lifting fan protection
        [0].rgxFault[0].4   // M310PopupUP.Lifting fan feedback
        [0].rgxWarning[0].0   // M310PopupUP.Positioning error on conveyor
        [1].rgxFault[0].0   // M310PopupDN.Lifting protection motor
        [1].rgxFault[0].1   // M310PopupDN.Lifting feedback motor
        [1].rgxFault[0].3   // M310PopupDN.Lifting fan protection
        [1].rgxFault[0].4   // M310PopupDN.Lifting fan feedback
        [1].rgxWarning[0].0   // M310PopupDN.Positioning error on conveyor
        [0].rgxStoppingFault[0].0   // M310PopupUP.Lifting position error
        [0].rgxFault[0].2   // M310PopupUP.Lifting safety switch
        [1].rgxStoppingFault[0].0   // M310PopupDN.Lifting position error
        [1].rgxFault[0].2   // M310PopupDN.Lifting safety switch
   M310Popup_HMR : MAC_Popup_ZC_HMR[2] := ([0].xHighPosition := 1, [0].rgdState := 1, [1].xHighPosition := 1, [1].rgdState := 1); {access Read Only}
        [0].rgxMan.0   // Rise popup upstream {x|x|x|x|O}
        [0].rgxMan.1   // Lower popup upstream {x|x|x|x|O}
        [0].rgxMan.2   // Rise both popup {x|x|x|x|O}
        [0].rgxMan.3   // Lower both popup {x|x|x|x|O}
        [1].rgxMan.0   // Rise popup downstream {x|x|x|x|O}
        [1].rgxMan.1   // Lower popup downstream {x|x|x|x|O}
   M310Popup_HMW : MAC_Popup_ZC_HMW[2] := ([0].dSingleCapOffset_cmm := 20000, [0].dSaturationSelection := 2);
        [0].rgxMan.0   // Rise popup upstream {x|x|x|x|O}
        [0].rgxMan.1   // Lower popup upstream {x|x|x|x|O}
        [0].rgxMan.2   // Rise both popup {x|x|x|x|O}
        [0].rgxMan.3   // Lower both popup {x|x|x|x|O}
        [1].rgxMan.0   // Rise popup downstream {x|x|x|x|O}
        [1].rgxMan.1   // Lower popup downstream {x|x|x|x|O}
   M310Popup_IN_MOTION : MAC_Popup_ZC_IN_MOTION[2]; {access None}
   M310Popup_OUT_MOTION : MAC_Popup_ZC_OUT_MOTION[2]; {access None}
   M310Popup_PlateFreeTimeout : TIMER; {access Read Only}
   M310Popup_ReentryCap : UDT_ConvoyCap_ZC;
   M310Popup_SL_DATA : UDT_Convoy_SL; {access Read Only}
   M310Popup_tSearchPlateChangeFromCS4401 : GP_TrackingSearchPlate_STC; {access Read Only}
   M310Popup_xDrivePosEnable : BOOL; {access Read Only}
   M310Popup_xEndRise : BOOL; {access Read Only}
   M310Popup_xEndRiseWaitingForCondition : BOOL; {access Read Only}
   M311 : MAC_Conveyor := (ST_xCleaningConditionOK := 1, ST_xEnableControlError := 1, ST_xPlateSynchronized := 1, ST_xSafetyMovement := 1, OSR_xSynchroPhotocellTail := 1, INPUT_xDriveReady_M1 := 1, INPUT_xLocalSafetySwitch_M1 := 1, INPUT_xMotorThermalProbe_M1 := 1, INPUT_xProtectionMotor_M1 := 1, INPUT_xDriveReady_M2 := 1, INPUT_xLocalSafetySwitch_M2 := 1, INPUT_xMotorThermalProbe_M2 := 1, INPUT_xProtectionMotor_M2 := 1, OUTPUT_xDriveEnable_M1 := 1, OUTPUT_xDriveEnable_M2 := 1, AUX_dPresetStopLoad_cmm := 408333, AUX_dPresetStopUnload_cmm := 491667, AUX_dAccSpace_cmm := 41667, AUX_dDecSpace_cmm := 41667, AUX_dReqSpeed_mm_min := 60000, AUX_dPhPosTarget_cmm := 295000, AUX_dPhPosTarget_2_cmm := 169750, tmON_FeedbackTimeOut_M1.PRE := 1500, tmOF_DriveEnable_M1.PRE := 30000, tmOF_DriveEnable_M1.ACC := 1820, tmOF_DriveEnable_M1.TT := 1, tmOF_DriveEnable_M1.DN := 1, tmOF_PowerSaving_M1.PRE := 20000, tmOF_PowerSaving_M1.ACC := 20000, tmON_FeedbackTimeOut_M2.PRE := 2000, tmOF_DriveEnable_M2.PRE := 30000, tmOF_DriveEnable_M2.ACC := 1820, tmOF_DriveEnable_M2.TT := 1, tmOF_DriveEnable_M2.DN := 1, tmOF_PowerSaving_M2.PRE := 20000, tmON_AuxFunction6.PRE := 5000, tmON_AuxFunction7.PRE := 100, tmON_AuxFunction8.PRE := 100, tmOF_MCD_M1.PRE := 200, tmOF_MCD_M1.ACC := 200, tmOF_MCD_M2.PRE := 200, tmOF_MCD_M2.ACC := 200); {access None}
        .INPUT_xMotorThermalProbe_M2   // M403.M2.P403BT4. Motor thermal probe
        .ST_xAux1   // request rise popup to unload on M325 (reentry)
        .INPUT_xMotorThermalProbe_M1   // M403.M1.P403BT3. Motor thermal probe
        .INPUT_xSyncroPhotocell_1   // M403.P115B1.Synchro photocell / start count
        .PH_x.0   // Load
        .PH_x.1   // Load Upstream
        .PH_x.10   // Unload Upstream
        .PH_x.11   // End load Downstream
        .PH_x.12   // Unload Downstream
        .PH_x.13   // End unload Upstream
        .PH_x.14   // End unload Downstream
        .PH_x.15   // End unload
        .PH_x.16   // Unload Unpack (n caps)
        .PH_x.17   // End unload Unpack (n caps)
        .PH_x.18   // Unload Unpack (n caps) Upstream
        .PH_x.19   // End unload Unpack (n caps) Upstream
        .PH_x.2   // Load Downstream
        .PH_x.20   // Unload Unpack (n caps) Downstream
        .PH_x.21   // End unload Unpack (n caps) Downstream
        .PH_x.22   // Load reentry
        .PH_x.23   // End load reentry
        .PH_x.24   // Unload reentry
        .PH_x.25   // End unload reentry
        .PH_x.26   // Load Unpack (n caps)
        .PH_x.27   // End load Unpack (n caps)
        .PH_x.28   // Load Unpack (n caps) Upstream
        .PH_x.29   // End load Unpack (n caps) Upstream
        .PH_x.3   // Wait rotation done
        .PH_x.30   // Load Unpack (n caps) Downstream
        .PH_x.31   // End load Unpack (n caps) Downstream
        .PH_x.4   // Rotation Ended
        .PH_x.7   // End load
        .PH_x.8   // Unload
        .PH_x.9   // End load Upstream
   M311_ALM : MAC_Conveyor_ALM;
        .rgdFaultCode_M[0]   // Drive fault code M1
        .rgdFaultCode_M[1]   // Drive fault code M2
        .rgxStoppingFault[0].0   // Z401.M311-M1.Positioning error
        .rgxStoppingFault[0].1   // Z401.M311-M1.Phase in progress with rotator not in low position
        .rgxStoppingFault_M[0].0   // Z401.M311-M1.Protection motor rotation
        .rgxStoppingFault_M[0].1   // Z401.M311-M1.Drive error
        .rgxStoppingFault_M[0].2   // Z401.M311-M1.Drive feedback error
        .rgxStoppingFault_M[0].3   // Z401.M311-M1.Local safety switch
        .rgxStoppingFault_M[0].4   // Z401.M311-M1.Motor thermal probe
        .rgxStoppingFault_M[0].5   // Z401.M311-M1.Braking resistor anomaly
        .rgxStoppingFault_M[0].6   // Z401.M311-M1.Drive not ready
        .rgxWarning[0].0   // Z401.M311.Plate not synchronized
        .rgxWarning[0].1   // Z401.M311.Positioning error
   M311_Data : UDT_Convoy_SL;
   M311_dLastRotationA_ID : DINT; {access Read Only}
   M311_HMR : MAC_Conveyor_HMR := (xIdPlatePresence := 1, dState1 := 1, dState2 := 1, dStateSensor1 := 1, dStateSensor2 := 1, dStateSensor3 := 1, dStateSensor4 := 1);
        .dErrorCode1   // Error code M1
        .rgxMan.0   // Run M1
        .rgxMan.1   // Reverse M1
        .rgxMan.2   // Run M2
        .rgxMan.3   // Reverse M2
